     ElseIf sender = 3 Then 'button "cut" is pressed
   	 If SmartTags("copyusb") = True Then
   		    SmartTags("AbufferFile") = SmartTags("File_"&SmartTags("fileChosen"))
   		    SmartTags("AbufferFolder") = SmartTags("Folder")
   		    SmartTags("AbufferCopyCut") = False 
   		    SmartTags("AbufferIsFolder") = SmartTags("isFolder_"&SmartTags("fileChosen"))
   		    SmartTags("AFEStatus") = "File " & SmartTags("AbufferFile") & " cut"
   	 Else    
   	   		SmartTags("AbufferFile") = SmartTags("aFile_"&SmartTags("AfileChosen"))
   		    SmartTags("AbufferFolder") = SmartTags("AFolder")
   		    SmartTags("AbufferCopyCut") = False 
   		    SmartTags("AbufferIsFolder") = SmartTags("aisFolder_"&SmartTags("AfileChosen"))
   		    SmartTags("AFEStatus") = "File " & SmartTags("AbufferFile") & " cut"
   	 End If  
     ElseIf sender = 2 Then 'button "move" pressed
       singleFile = Replace (SmartTags("AbufferFile"),  SmartTags("AbufferFolder"), "")
       newpath = SmartTags("AFolder") & singleFile  
       If SmartTags("AbufferCopyCut") = False Then   
         If SmartTags("AbufferIsFolder") <> 0 Then
           Set fs = CreateObject("FileCtl.FileSystem")
           fs.MoveFile SmartTags("AbufferFile"), newpath
         Else
           Set fs = CreateObject("FileCtl.FileSystem")
           fs.FileCopy SmartTags("AbufferFile"), newpath
           fs.kill SmartTags("AbufferFile")
         End If
       Else
         Set fs = CreateObject("FileCtl.FileSystem")
         fs.FileCopy SmartTags("AbufferFile"), newpath
       End If 
       SmartTags("AFEStatus") = "File " & SmartTags("AbufferFile") & " pasted"
       LHmiView_vbsFEReadFilesOfFolder_1 SmartTags("AFolder")
       LHmiView_vbsFEWriteFilePropertiesToTags_1 SmartTags("Aindex")
     End If
   ' Windows / PC based
   Else
     If sender = 1 Then 'button "copy" pressed
   	  'edit agar dapat copy local dir / external dir
   	  If SmartTags("copyusb") = True Then 
       	SmartTags("AbufferFile") = SmartTags("File_"&SmartTags("fileChosen"))
      		SmartTags("AbufferFolder") = SmartTags("Folder")
       	SmartTags("AbufferCopyCut") = True
       	SmartTags("AbufferIsFolder") = SmartTags("isFolder_"&SmartTags("fileChosen"))
       	SmartTags("AFEStatus") = "File " & SmartTags("AbufferFile") & " copied"
   	  Else
   		SmartTags("AbufferFile") = SmartTags("aFile_"&SmartTags("AfileChosen"))
      		SmartTags("AbufferFolder") = SmartTags("AFolder")
       	SmartTags("AbufferCopyCut") = True
       	SmartTags("AbufferIsFolder") = SmartTags("aisFolder_"&SmartTags("AfileChosen"))
       	SmartTags("AFEStatus") = "File " & SmartTags("AbufferFile") & " copied" 
   	  End If
   	  
     ElseIf sender = 3 Then 'button "cut" is pressed
        'edit agar dapat copy local dir / external dir
        If SmartTags("copyusb") = True Then 
      		SmartTags("AbufferFile") = SmartTags("File_"&SmartTags("fileChosen"))
     		SmartTags("AbufferFolder") = SmartTags("Folder")
       	SmartTags("AbufferCopyCut") = False 
   		SmartTags("AbufferIsFolder") = SmartTags("isFolder_"&SmartTags("fileChosen"))
   		SmartTags("AFEStatus") = "File " & SmartTags("AbufferFile") & " cut"
   	 Else
   		 SmartTags("AbufferFile") = SmartTags("aFile_"&SmartTags("AfileChosen"))
      		 SmartTags("AbufferFolder") = SmartTags("AFolder")
      		 SmartTags("AbufferCopyCut") = False 
      		 SmartTags("AbufferIsFolder") = SmartTags("aisFolder_"&SmartTags("AfileChosen"))
       	 SmartTags("AFEStatus") = "File " & SmartTags("AbufferFile") & " cut"
       End If
       
     ElseIf sender = 2 Then 'button "move" pressed
       singleFile = Replace (SmartTags("AbufferFile"),  SmartTags("AbufferFolder"), "")
       newpath = SmartTags("AFolder") & singleFile  
       Set fs = CreateObject("Scripting.FileSystemObject")
       If SmartTags("AbufferCopyCut") = False Then
         If SmartTags("AbufferIsFolder") = "True" Then
           data = fs.GetFolder(SmartTags("AbufferFile"))
           fs.MoveFolder data, newpath
         Else
           data = fs.GetFile(SmartTags("AbufferFile"))
           fs.MoveFile data, newpath
         End If
       Else
         If SmartTags("AbufferIsFolder") = "True" Then
           data = fs.GetFolder(SmartTags("AbufferFile"))
           fs.CopyFolder data, newpath
         Else
           data = fs.GetFile(SmartTags("AbufferFile"))
           fs.CopyFile data, newpath
         End If
       End If
       If Err.Number <> 0 Then
         SmartTags("AFEStatus") = Err.Description & "Could not paste file / folder"
       Else
         SmartTags("AFEStatus") = "File / Folder " & SmartTags("AbufferFile") & " pasted"
       End If
       LHmiView_vbsFEReadFilesOfFolder_1 SmartTags("AFolder")
       LHmiView_vbsFEWriteFilePropertiesToTags_1 SmartTags("Aindex")
     End If
   End If

VB script "LHmiView_vbsFEDelete_1"
   On Error Resume Next
   
   '-----------------------DEFINE PARAMETERS-------------------------------------------
   'kindOfOperatingSystem: 0 = Windows, 1 = Windows CE
   ' tempFs: Reference on temporary fileSystem Object
   ' fs: Reference on fileSystem Object
   ' f: Reference on file Object
   Dim kindOfOperatingSystem, tempFs, f, fs, file
   
   '--------------------Prove which Operating System is running------------------------
   'Set tempFs = CreateObject("Scripting.FileSystemObject")
   
   'If Err.Number = 0 Then
   '	kindOfOperatingSystem = 0 'Windows / PC based
   'Else
   	kindOfOperatingSystem = 1 'Windows CE / Panel based
   'End If
   
   Set tempFs= Nothing
   Err.Clear
   
   '-------------------------------Delete folder/file---------------------------------
   Dim i
   
   SmartTags("AFEStatus") = "Deleting file..."
   i = SmartTags("AfileChosen")
   
   ' Windows CE / Panel based
   If kindOfOperatingSystem Then    
     Set fs = CreateObject("FileCtl.FileSystem")
     Set f = CreateObject("FileCtl.File")
     If i > 0 And SmartTags("aFile_"&i) <> "" Then
       If SmartTags("aisFolder_"&i) <> 0 Then
         fs.RmDir SmartTags("aFile_"&i)
         If Err.Number = 0 Then
           SmartTags("AFEStatus") = "File / Folder deleted: " & SmartTags("aFile_"&i) 
           SmartTags("aFile_"&i) = ""
         Else
           SmartTags("AFEStatus") = "Could not delete file / folder: " & SmartTags("aFile_"&i)
         End If
       Else
         fs.kill SmartTags("aFile_"&i)
         If Err.Number = 0 Then
           SmartTags("AFEStatus") = "File / Folder deleted: " & SmartTags("aFile_"&i) 
         Else
           SmartTags("AFEStatus") = "Could not delete file / folder: " & SmartTags("aFile_"&i)
         End If
         SmartTags("aFile_"&i) = ""
       End If
     Else
       SmartTags("AFEStatus") = "Choose file / folder"
     End If
     
   ' Windows / PC based
   Else
     Set fs = CreateObject("Scripting.FileSystemObject")
      If i > 0 And SmartTags("aFile_"&i) <> "" Then
       If SmartTags("aisFolder_"&i) <> "False" Then
         fs.DeleteFolder(SmartTags("aFile_"&i))
         If Err.Number = 0 Then
           SmartTags("AFEStatus") = "File / folder deleted: " & SmartTags("aFile_"&i) 
           SmartTags("aFile_"&i) = ""
         Else
           SmartTags("AFEStatus") = "Could not delete file / folder: " & SmartTags("aFile_"&i)
         End If
       Else
         fs.DeleteFile(SmartTags("aFile_"&i))
         If Err.Number = 0 Then
           SmartTags("AFEStatus") = "Folder / folder deleted: " & SmartTags("aFile_"&i) 
         Else
           SmartTags("AFEStatus") = "Could not delete file/ folder: " & SmartTags("aFile_"&i)
         End If
         SmartTags("aFile_"&i) = ""
       End If
     Else
       SmartTags("AFEStatus") = "Choose file / folder"
     End If
   End If
   
   Set fs = Nothing
   Set f = Nothing
   
   LHmiView_vbsFEReadFilesOfFolder_1 SmartTags("AFolder")
   LHmiView_vbsFEWriteFilePropertiesToTags_1 SmartTags("Aindex")

VB script "delfunc"
   Dim i
   
   For i= 1 To 10
   	SmartTags("AisFolder_" &i) = 0
   Next

VB script "Delay"
   Dim StartTime, StopTime, i , x
   
   StartTime = Now
   StopTime = Now + DelayTime/3600/154
   
   Do
   Loop Until Now >= StopTime

scheduled task "User_Change"
   on Action: function_e1ab61de("NavUserChange")
*)